VAR_GLOBAL CONSTANT   // PLC tag table "STEP7 classic symbols"
   "A" : Real := 0.5485;
   "B" : Real := 0.665E-3;
   "C" : Real := 2.805E-9;
   "A_FC343" : Real := 3.90802E-3;   // MigChange: A
   "B_FC343" : Real := -5.802000E-007;   // MigChange: B , -5.802E-7
   "C_FC343" : Real := -4.273500E-012;   // MigChange: C , -4.27350E-12
   "A_FC344" : Real := 7.64E-3;   // MigChange: A
   "B_FC344" : Real := 1.66E-5;   // MigChange: B
   "A_FC347" : Real := 3.9083E-3;   // MigChange: A
   "B_FC347" : Real := -5.775000E-007;   // MigChange: B , -5.775E-7
   "accuracy" : Real := 0.01;
END_VAR

FUNCTION "MID3" : Real   // FC96, SCL
TITLE = MID3
{ S7_Optimized_Access := 'FALSE' }
AUTHOR : hugo
FAMILY : MATH
NAME : MID3
VERSION : 1.2
// returns the mid value of 3 real inputs.
   VAR_INPUT
      in1 : Real;
      in2 : Real;
      in3 : Real;
   END_VAR
   VAR_TEMP
      tIN1 : Real;
      tIN2 : Real;
      tIN3 : Real;
   END_VAR
BEGIN


   #tIN1 := #in1;
   #tIN2 := #in2;
   #tIN3 := #in3;

   IF #tIN1 > #tIN2 THEN 
     #MID3 := #tIN1; 
     #tIN1 := #tIN2; 
     #tIN2 := #MID3; 
   END_IF;

   IF #tIN2 > #tIN3 THEN 
     #tIN2 := #tIN3; 
   END_IF;

   #MID3 := SEL(G:=#tIN1 > #tIN2, IN0:=#tIN2, IN1:=#tIN1);

   (*
   hm  1.1.2007  rev 1.1
     rewrote the function for better performance

   hm  18. mar. 2011 rev 1.2
     improve performance
   *)
END_FUNCTION

FUNCTION "MULTI_IN" : Real   // FC341, SCL
TITLE = MULTI_IN
{ S7_Optimized_Access := 'FALSE' }
AUTHOR : oscat
FAMILY : SENSOR
NAME : MULTI_IN
VERSION : 1.4
// multi_in is a signal conditioning function ehich can be configured in 8 different ways.
// it is used to read multiple sensors for the same value and protect the user from broken sensors or invalid data from sensors.
//  
// multi_in can be configured in different ways:
//     mode = 0 means the the avg of the 3 inputs is used, this mode is the default mode.
//     mode = 1 means in_1 is used.
//     mode = 2 means in_2 is used.
//     mode = 3 means in_3 is used.
//     mode = 4 means default is used.
//     mode = 5 means the lowest of the 3 external temperatures is used.
//     mode = 6 means the higest externnal temperature is used.
//     mode = 7 means the midlle input is used, if there are only two working, the lowest input is used.
//     mode > 7 ,eans output is 0 at all times.
//     in any config mode, an input higher then in_max or lower then in_min is ignored to prevent values from broken sensors or wires.
//     if all inputs are higher then in_max or lower then in_min, a default value (default) is used.
// 
// uses: MID3 [FC96]
   VAR_INPUT
      in_1 : Real;
      in_2 : Real;
      in_3 : Real;
      default : Real;
      in_min : Real;
      in_max : Real;
      mode : Int;
   END_VAR
   VAR_TEMP
      count : Int;
      F1 : Bool;
      F2 : Bool;
      F3 : Bool;
   END_VAR
BEGIN


   #F1 :=  #in_1 > #in_min AND #in_1 < #in_max;
   #F2 :=  #in_2 > #in_min AND #in_2 < #in_max;
   #F3 :=  #in_3 > #in_min AND #in_3 < #in_max;

   CASE #mode OF
   0:  #count := 0;
     IF #F1 THEN
       #count := #count + 1;
       #MULTI_IN := #in_1;
     ELSE
       #MULTI_IN := 0.0;
     END_IF;
     IF #F2 THEN
       #count := #count + 1;
       #MULTI_IN := #MULTI_IN + #in_2;
     END_IF;
     IF #F3 THEN
       #count := #count + 1;
       #MULTI_IN := #MULTI_IN + #in_3;
     END_IF;
     #MULTI_IN := SEL(G:=#count = 0, IN0:=#MULTI_IN / INT_TO_REAL(#count), IN1:=#default);

   1:  #MULTI_IN := SEL(G:=#F1, IN0:=#default, IN1:=#in_1);

   2:  #MULTI_IN := SEL(G:=#F2, IN0:=#default, IN1:=#in_2);

   3:  #MULTI_IN := SEL(G:=#F3, IN0:=#default, IN1:=#in_3);

   4:  #MULTI_IN := #default;

   5:  #MULTI_IN := SEL(G:=#F1, IN0:=#in_max, IN1:=#in_1);
     IF #F2 AND #in_2 < #MULTI_IN THEN #MULTI_IN := #in_2; END_IF;
     IF #F3 AND #in_3 < #MULTI_IN THEN #MULTI_IN := #in_3; END_IF;
     IF #MULTI_IN = #in_max THEN #MULTI_IN := #default; END_IF;

   6:  #MULTI_IN := SEL(G:=#F1, IN0:=#in_min, IN1:=#in_1);
     IF #F2 AND #in_2 > #MULTI_IN THEN #MULTI_IN := #in_2; END_IF;
     IF #F3 AND #in_3 > #MULTI_IN THEN #MULTI_IN := #in_3; END_IF;
     IF #MULTI_IN = #in_min THEN #MULTI_IN := #default; END_IF;

   7:  IF #F1 AND #F2 AND #F3 THEN #MULTI_IN := "MID3"(in1:=#in_1, in2:=#in_2, in3:=#in_3);
     ELSIF #F1 AND #F2 THEN #MULTI_IN := MIN(IN1:=#in_1, IN2:=#in_2);
     ELSIF #F1 AND #F3 THEN #MULTI_IN := MIN(IN1:=#in_1, IN2:=#in_3);
     ELSIF #F2 AND #F3 THEN #MULTI_IN := MIN(IN1:=#in_2, IN2:=#in_3);
     ELSIF #F1 THEN #MULTI_IN := #in_1;
     ELSIF #F2 THEN #MULTI_IN := #in_2;
     ELSIF #F3 THEN #MULTI_IN := #in_3;
     ELSE #MULTI_IN := #default;
     END_IF;

   END_CASE;

   (*
   hm 1.1.2007   rev 1.1
     changed midr to mid3 function

   hm  14. 10. 2008  rev 1.2
     corrected an error for in_3 overrange detection
     improved performance

   hm  11. mar. 2009 rev 1.3
     changed real constants to use dot syntax

   hm  18. jul. 2009 rev 1.4
     improved performance
   *)
END_FUNCTION

FUNCTION "RES_NI" : Real   // FC342, SCL
TITLE = RES_NI
{ S7_Optimized_Access := 'FALSE' }
AUTHOR : hugo
FAMILY : SENSOR
NAME : RES_NI
VERSION : 1.2
// this function returs the resistance for a nickel sensor for a temperature range from -60..+180 °C
   VAR_INPUT
      T : Real;
      R0 : Real;
   END_VAR
   VAR_TEMP
      T_2 : Real;
   END_VAR
BEGIN


     #T_2 := #T*#T;
     #RES_NI := #R0 + "A"*#T + "B"*#T_2 + "C"*#T_2*#T_2;


   (* revision history

   hm  4.8.2006    rev 1.0
     original version

   hm  13.9.2007    rev 1.1
     changed coding for better performance

   hm  2. dec. 2007  rev 1.2
     changed code for better performance
   *)

   (*

    Auszug aus DIN 43760 für Ni100

   °C    R    °C    R    °C  R    °C    R    °C    R

   -60   69,5   -10   94,6   40   123,0   90     154,9   140   190,9
   -55   71,9   -5     97,3   45   126,0   95     158,3   145   194,8
   -50   74,3   0     100,0   50   129,1   100   161,8   150   198,7
   -45   76,7   5     102,8   55   132,2   105   165,3   155   202,6
   -40   79,1   10     105,6   60   135,3   110   168,8   160   206,6
   -35   81,6   15     108,4   65   138,5   115   172,4   165   210,7
   -30   84,2   20     111,2   70   141,7   120   176,0   170   214,8
   -25   86,7   25     114,1   75   145,0   125   179,6   175   219,0
   -20   89,3   30     117,1   80   148,3   130   183,3   180   223,2
   -15   91,9   35     120,0   85   151,6   135   187,1        

   *)
END_FUNCTION

FUNCTION "RES_PT" : Real   // FC343, SCL
TITLE = RES_PT
{ S7_Optimized_Access := 'FALSE' }
AUTHOR : hugo
FAMILY : SENSOR
NAME : RES_PT
VERSION : 1.3
// this function returs the resistance for a platinum sensor for a temperature range from -200..+850 °C
   VAR_INPUT
      T : Real;
      R0 : Real;
   END_VAR
   VAR_TEMP
      T_2 : Real;
   END_VAR
BEGIN


   #T_2 := #T * #T;

   IF #T >= 0.0 THEN
       #RES_PT := #R0 * ( 1.0 + "A"* #T + "B_FC343" * #T_2);
   ELSE
       #RES_PT := #R0 * ( 1.0 + "A"* #T + "B_FC343" * #T_2 + "C_FC343" *(#T - 100.0) * #T_2 * #T);
   END_IF;


   (* revision history
   hm  4. aug. 2006    rev 1.1
       original version

   hm  2. dec 2007 rev 1.2
       changed code for better performance

   hm  11. mar. 2009   rev 1.3
       changed real constants to use dot syntax

   *)


   (*
    Auszug aus DIN 43760 für Pt100

   °C      R       °C      R       °C  R           °C      R           °C      R           °C      R

   -200    18,49   -100    60,25   0   100,00  100     138,50  200     175,84  300     212,02
   -195    20,65   -95     62,28   5   101,95  105     140,39  205     177,68  305     213,80
   -190    22,80   -90     64,30   10  103,90  110     142,29  210     179,51  310     215,57
   -185    24,94   -85     66,31   15  105,85  115     144,17  215     181,34  315     217,35
   -180    27,08   -80     68,33   20  107,79  120     146,06  220     183,17  320     219,12
   -175    29,20   -75     70,33   25  109,73  125     147,94  225     184,99  325     220,88
   -170    31,32   -70     72,33   30  111,67  130     149,82  230     186,82  330     222,65
   -165    33,43   -65     74,33   35  113,61   135     151,70  235     188,63  335     224,41
   -160    35,33   -60     76,33   40  115,54  140     153,58  240     190,45  340     226,17
   -155    37,63   -55     78,32   45  117,47  145     155,45  245     192,26  345     227,92
   -150    39,71   -50     80,31   50  119,40  150     157,31  250     194,07  350     229,67
   -145    41,79   -45     82,29   55  121,32  155     159,18  255     195,88  355     231,42
   -140    43,87   -40     84,27   60  123,24  160     161,04  260     197,69  360     233,17
   -135    45,94   -35     86,25   65  125,16  165     162,90  265     199,49  365     234,91
   -130    48,00  -30     88,22   70  127,07  170     164,76  270     201,29  370     236,65
   -125    50,06   -25     90,19   75  128,98  175     166,61  275     203,08  375     238,39
   -120    52,11   -20     92,16   80  130,89  180     168,46  280     204,88  380     240,13
   -115    54,15   -15     94,12   85  132,80  185     170,31  285     206,67  385     241,86
   -110    56,19   -10     96,09   90  134,70  190     172,16  290     208,45  390     243,59
   -105    58,22   -5      98,04   95  136,60  195     174,00  295     210,24  395     245,31

   *)
   (*
   revision history


   *)
END_FUNCTION

FUNCTION "RES_SI" : Real   // FC344, SCL
TITLE = RES_SI
{ S7_Optimized_Access := 'FALSE' }
AUTHOR : hugo
FAMILY : SENSOR
NAME : RES_SI
VERSION : 1.2
// this function returs the resistance for a silicon sensor for a temperature range from -50..+150 °C
// for example KTY10 normaly Rs at 25 °C
   VAR_INPUT
      T : Real;
      RS : Real;
      TS : Real;
   END_VAR
   VAR_TEMP
      TX : Real;
   END_VAR
BEGIN


   #TX := #T - #TS;
   #RES_SI := #RS * ( 1.0 + "A"* #TX + "B_FC344" * #TX * #TX);


   (* revision history
   hm  4. aug 2006 rev 1.0
       original version

   hm  2. dec 2007 rev 1.1
       changed code for better performance

   hm  11. mar. 2009   rev 1.2
       changed real constants to use dot syntax

   *)
END_FUNCTION

FUNCTION "SENSOR_INT" : Real   // FC345, SCL
TITLE = SENSOR_INT
{ S7_Optimized_Access := 'FALSE' }
AUTHOR : hugo
FAMILY : SENSOR
NAME : SENS_INT
VERSION : 1.3
// this FUNCTION calculates the REAL resistance OF a sensor RX given a parasitic resistor in parallel TO the sensor AND an additional serial resistor.
// for example a parasitic parallel resistor for a PT100 can be ignored but a series resistor is the cable to the sensor.
// for a humidity sensor, the parallel resistor is more dramatic and needs to be considered.
// the function allows to consider a parallel and serial resistor at the same time.
// with this function and known parasitic serial and parallel resistors the true resistance of the sensor can be calculated.
   VAR_INPUT
      Voltage : Real;
      Current : Real;
      RP : Real;
      RS : Real;
   END_VAR
   VAR_TEMP
      RG : Real;
   END_VAR
BEGIN


   IF #Current <> 0.0 THEN
       #RG := #Voltage / #Current;
       #SENSOR_INT := #RP * ( #RG - #RS) / ( #RP + #RS - #RG);
   END_IF;


   (* revisaion history

   hm 20.1.2007        rev 1.1
       deleted input R0 which was not needed.

   hm  2. dec 2007 rev 1.2
       corrected an error in formula and improoved speed

   hm  11. mar. 2009   rev 1.3
       changed real constants to use dot syntax

   *)
END_FUNCTION

FUNCTION "TEMP_NI" : Real   // FC346, SCL
TITLE = TEMP_NI
{ S7_Optimized_Access := 'FALSE' }
AUTHOR : hugo
FAMILY : SENSOR
NAME : TEMP_NI
VERSION : 1.5
// this function returs the temperature for a nickel sensor for a range from -60..+180 °C
   VAR_INPUT
      Res : Real;
      R0 : Real;
   END_VAR
BEGIN


   #TEMP_NI := (SQRT(0.30085225 - 2.66E-3 * (#R0 - #Res)) - 0.5485) * 751.8796992;


   (* revision history

   hm 24.1.2007        rev 1.1
       deleted unused variable A, B, C

   hm 10.9.2007        rev 1.2
       changed accuracy to 0.02 degrees to improove performace

   hm 17. 12 2007  rev 1.3
       improovements for better performance and higher accuracy

   hm  6. jan 2008 rev 1.4
       further performance improvement

   hm  10. mar. 2009   rev 1.5
       removed nested comments

   *)
END_FUNCTION

FUNCTION "TEMP_PT" : Real   // FC347, SCL
TITLE = TEMP_PT
{ S7_Optimized_Access := 'FALSE' }
AUTHOR : hugo
FAMILY : SENSOR
NAME : TEMP_PT
VERSION : 1.7
// this function returs the temperature for a platinum sensor for a range from -200..+850 °C 
// 
// uses: RES_PT [FC343]
   VAR_INPUT
      Res : Real;
      R0 : Real;
   END_VAR
   VAR_TEMP
      "step" : Real;
      X : Real;
      Y : Real;
      t1 : Real;
   END_VAR
BEGIN


   #"step" := 50.0;

   #X := "A"* #R0;
   #Y := "B_FC347" * #R0;
   IF #Res >= #R0 THEN
       #t1 := #X * #X - 4.0 * #Y * (#R0 - #Res);
       IF #t1 < 0.0 THEN
           #TEMP_PT := 10000.0;
       ELSE
           #TEMP_PT := (-#X + SQRT(#t1)) / (2.0 * #Y);
       END_IF;
   ELSE
       (* since the formula cannot be solved this is a successive approximation *)
       #TEMP_PT := -100.0;
       WHILE #"step" > "accuracy" DO
           (* test if result greater or less *)
           IF "RES_PT"(T:=#TEMP_PT,R0:=#R0) < #Res THEN #TEMP_PT := #TEMP_PT + #"step"; ELSE #TEMP_PT := #TEMP_PT - #"step"; END_IF;
           (* pt^ := pt^ - 8388608; *)  (* this is a super fast divide by 2 method for non floating point CPUs *)
           (* the alternative code: step := step * 0.5; *)
           #"step" := #"step" * 0.5;
       END_WHILE;
   END_IF;

   (* revision history

   rev 1.1 hm 24.1.2007    
       deleted unused variable C

   rev 1.2 hm 10.9.2007
       reduced accuracy to 0.02 to shorten execution time

   rev 1.3 hm  2. dec 2007
       changed code for better performance

   rev 1.4 hm  23. dec 2007
       avoid a negative square root if input values are wrong

   rev 1.5 hm 5. jan 2008
       replaced / 2 with * 0.5 for better performance

   hm  31. oct. 2008   rev 1.6
       improved performance

   hm  11. mar. 2009   rev 1.7
       changed real constants to use dot syntax

   *)
END_FUNCTION

FUNCTION "TEMP_SI" : Real   // FC348, SCL
TITLE = TEMP_SI
{ S7_Optimized_Access := 'FALSE' }
AUTHOR : hugo
FAMILY : SENSOR
NAME : TEMP_SI
VERSION : 1.5
// this function returs the temperature for a silicon sensor for a range from -50..+150 °C
// for example KTY10 RS at TS normally 25 °C
   VAR_INPUT
      Res : Real;
      RS : Real;
      TS : Real;
   END_VAR
BEGIN


   #TEMP_SI := (-7.64E-3 + SQRT(#Res/#RS* 6.64E-5 - 0.803E-5)) * 30120.48193 + #TS;


   (* revision history

   hm 24.1.2007        rev 1.1
       the function would only work for TS = 25, now it works for other values of ts.

   hm 10.9.2007        rev 1.2
       changed the function to use successive approcimation to avoid an error generated by a sqrt from a negative result.
       changed accuracy to 0.02 degrees to shorten execution time

   hm 17. 12 2007  rev 1.3
       improovements for better performance

   hm  6. jan 2008 rev 1.4
       further performance improvement

   hm  10. mar. 2009   rev 1.5
       removed nested comments

   *)
END_FUNCTION

FUNCTION "TEMP_NTC" : Real   // FC411, SCL
TITLE = TEMP_NTC
{ S7_Optimized_Access := 'FALSE' }
AUTHOR : hugo
FAMILY : SENSOR
NAME : TEMP_NTC
VERSION : 1.1
// this function returs the temperature for a NTC sensor for a range from 0..85 °C.
// RN is the resistance at 25 °C and B is a constant for the given sensor.
   VAR_INPUT
      RES : Real;
      RN : Real;
      "B" : Real;
   END_VAR
BEGIN


   IF #RES > 0.0 THEN
       #TEMP_NTC := #"B" * 298.15 / (#"B" + LN(#RES / #RN) * 298.15) -273.15;
   END_IF;


   (* revision history

   hm 30. dec. 2008    rev 1.0
       original version

   hm  11. mar. 2009   rev 1.1
       changed real constants to use dot syntax

   *)
END_FUNCTION

FUNCTION "RES_NTC" : Real   // FC412, SCL
TITLE = RES_NTC
{ S7_Optimized_Access := 'FALSE' }
AUTHOR : hugo
FAMILY : SENSOR
NAME : RES_NTC
VERSION : 1.1
// this function returs the resistance for a NTC sensor for a given temperature in °C.
// RN is the resistance at 25 °C and B is a constant for the given sensor.
   VAR_INPUT
      T : Real;
      RN : Real;
      "B" : Real;
   END_VAR
BEGIN


   #RES_NTC := #RN * EXP(#"B" * (1.0 / (#T+273.15) - 0.00335401643468053));


   (* revision history

   hm 30. dec. 2008    rev 1.0
       original version

   hm  11. mar. 2009   rev 1.1
       changed real constants to use dot syntax

   *)
END_FUNCTION

// ===== PLC "List Processing"  Unspecific CPU S7 300 =====

DATA_BLOCK "TEMP"   // DB7
TITLE = temporary Strings
{ S7_Optimized_Access := 'FALSE' }
AUTHOR : dalbi
FAMILY : xS7
NAME : DBTEMP
VERSION : 1.1
   VAR
      STR1 : String[254];
      STR2 : String[254];
      STR3 : String[254];
      TEMP : String[254];
   END_VAR
BEGIN
END_DATA_BLOCK

FUNCTION_BLOCK "LIST_NEXT"   // FB231, SCL
TITLE = LIST_NEXT
{ S7_Optimized_Access := 'FALSE' }
AUTHOR : hugo
FAMILY : LISTPRO
NAME : LNEXT
VERSION : 2.0
// LIST_NEXT retrieves the next element of a list, starting from element 1 after reset or first init.
// when the end of the lisat is reached a '' empty string is returned and NUL is set to true.
// die liste liegt als string von elementen vor die mit den zeichen SEP am anfang markiert sind.
   VAR_INPUT
      SEP : Byte;
      RST : Bool;
   END_VAR
   VAR_OUTPUT
      LEL : String[254];
      po AT LEL : Struct
         length : Byte;
         act_length : Byte;
         str : Array[1..254] of Byte;
      END_STRUCT;
      NUL : Bool;
   END_VAR
   VAR_IN_OUT
      LIST : String[254];
      pt AT LIST : Struct
         length : Byte;
         act_length : Byte;
         str : Array[1..254] of Byte;
      END_STRUCT;
   END_VAR
   VAR
      pos : Int := 1;
      c : Byte;
      write : Int;
   END_VAR
BEGIN


   //pt := ADR(LIST);
   //po := ADR(LEL);

   IF #RST THEN
     #pos := 1;
   END_IF;

   IF #pt.str[#pos] = 0 OR #pos = BYTE_TO_INT(#pt.act_length) THEN
     #LEL := '';
     #NUL := TRUE;
   ELSE
     #NUL := FALSE;
     #write := 1;
     FOR #pos := #pos + 1 TO BYTE_TO_INT(#pt.act_length) DO
       #c := #pt.str[#pos];
       IF #c = 0 OR #c = #SEP THEN
         #po.str[#write] := 0;
         RETURN;
       ELSE
         #po.str[#write] := #pt.str[#pos];
         #write := #write + 1;
       END_IF;
     END_FOR;
   END_IF;

   #po.length := #pt.length;
   #po.act_length := INT_TO_BYTE(#write);


   (* revision histroy
   hm  25. jun. 2008 rev 1.0
     original release

   hm  19. jan. 2011 rev 1.1
     changed string(255) to string(LIST_LENGTH)  

   hm  21. mar. 2011 rev 2.0
     all elements start with SEP

   *)
END_FUNCTION_BLOCK

FUNCTION "CHR_TO_STRING" : String[254]   // FC227, SCL
TITLE = CHR_TO_STRING
{ S7_Optimized_Access := 'FALSE' }
AUTHOR : hugo
FAMILY : STRINGS
NAME : CHRSTR
VERSION : 1.3
// CHR creates a character from a byte input and stuffs it in a one character length string.
   VAR_INPUT
      C : Byte;
   END_VAR
   VAR_TEMP
      tCHR : String[1];
      _CHR AT tCHR : Array[0..2] of Byte;
   END_VAR
BEGIN


   #_CHR[0] := 1;   (* length *)
   #_CHR[1] := 1;   (* actual length *)
   #_CHR[2] := #C; 
   #CHR_TO_STRING := #tCHR;

   (* revision history
   hm  16 jan 2007     rev 1.0
       original version

   hm  4. feb. 2008    rev 1.1
       return string would not be terminated properly

   hm  29. mar. 2008   rev 1.2
       changed STRING to STRING(1)

   hm  17. dec. 2008   rev 1.3
       changed name of function from chr to chr_to_string
   *)
END_FUNCTION

FUNCTION "LIST_CLEAN" : Bool   // FC389, SCL
TITLE = LIST_CLEAN
{ S7_Optimized_Access := 'FALSE' }
AUTHOR : hugo
FAMILY : LISTPRO
NAME : LCLEAN
VERSION : 2.0
// LIST_CLEAN bereinigt eine liste von leeren Elementen.
// die liste liegt als string von elementen vor die mit den zeichen SEP am anfang markiert sind.
   VAR_INPUT
      SEP : Byte;
   END_VAR
   VAR_IN_OUT
      LIST : String[254];
      pt AT LIST : Struct
         length : Byte;
         act_length : Byte;
         str : Array[1..254] of Byte;
      END_STRUCT;
   END_VAR
   VAR_TEMP
      read : Int;
      write : Int;
      last : Byte;
      c : Byte;
   END_VAR
BEGIN


   #read := 1;
   #write := 1;

   FOR #read := 1 TO BYTE_TO_INT(#pt.act_length) DO //LIST_LENGTH = 254
     #c := #pt.str[#read];               (* read character from list *)
     IF #c = 0 THEN EXIT;           (* exit the loop if character definbes end of string *)
     ELSIF #c <> #SEP OR #SEP <> #last THEN  (* copy element from read to write position unless a double sep character is present *)
       #pt.str[#write] := #c;
       #write := #write + 1;
     END_IF;
     #last := #c;                  (* remember last character *)
   END_FOR;

   IF #last = #SEP THEN #write := #write - 1; END_IF;    (* if last character is sep then delete empty element at end *)
   IF #write <= BYTE_TO_INT(#pt.act_length) THEN #pt.str[#write] := 0;  END_IF;    (* terminate string with 0 *)

   #LIST_CLEAN := TRUE;           (* retrun TRUE *)


   (* revision histroy
   hm  28. jun. 2008 rev 1.0
     original release

   hm  19. jan. 2011 rev 1.1
     changed string(255) to string(LIST_LENGTH)

   hm  21. mar. 2011 rev 2.0
     all elements start with SEP

   *)
END_FUNCTION

FUNCTION "LIST_GET" : String[254]   // FC390, SCL
TITLE = LIST_GET
{ S7_Optimized_Access := 'FALSE' }
AUTHOR : hugo
FAMILY : LISTPRO
NAME : LGET
VERSION : 2.0
// LIST_GET liefert das element an der stelle pos einer liste.
// die liste liegt als string von elementen vor die mit den zeichen SEP am anfang makiert sind.
   VAR_INPUT
      SEP : Byte;
      POS : Int;
   END_VAR
   VAR_IN_OUT
      LIST : String[254];
      pt AT LIST : Struct
         length : Byte;
         act_length : Byte;
         str : Array[1..254] of Byte;
      END_STRUCT;
   END_VAR
   VAR_TEMP
      tLIST_GET : String[254];
      po AT tLIST_GET : Struct
         length : Byte;
         act_length : Byte;
         str : Array[1..254] of Byte;
      END_STRUCT;
      i : Int;
      o : Int;
      cnt : Int;
      c : Byte;
   END_VAR
BEGIN


   #i := 1;
   #o := 1;
   #cnt := 0;

   REPEAT
     #c := #pt.str[#i];
     IF #cnt = #POS THEN           (* copy element to output string *)
       IF #c = #SEP  THEN EXIT; END_IF;    (* next element stop copy and finish *)
       #po.str[#o] := #c;
       #o := #o + 1;
     ELSIF #c = #SEP THEN
       #cnt := #cnt + 1;
     END_IF;
     #i := #i + 1;
   UNTIL
     (#i = BYTE_TO_INT(#pt.act_length)) OR (#c = 0)
   END_REPEAT;
   #po.act_length := INT_TO_BYTE(#o);            (* close the output string *)
   #po.length := #pt.length;

   #LIST_GET := #tLIST_GET;


   (* revision histroy
   hm  20. jun. 2008 rev 1.0
     original release

   hm  19. jan. 2011 rev 1.1
     changed string(255) to strring(LIST_LENGTH)

   hm  21. mar. 2011 rev 2.0
     all list elements start with SEP
   *)
END_FUNCTION

FUNCTION "LIST_INSERT" : Bool   // FC391, SCL
TITLE = LIST_INSERT
{ S7_Optimized_Access := 'FALSE' }
AUTHOR : hugo
FAMILY : LISTPRO
NAME : LINS
VERSION : 2.0
// LIST_INSERT setzt ein element an der stelle pos in eine liste ein.
// die liste liegt als string von elementen vor die mit den zeichen SEP am anfang markiert sind.
// 
// uses: CONCAT [FC2]
//       CHR_TO_STRING [FC227]
//       INSERT [FC17]
//       LEN [FC21]
//       TEMP [DB7]
   VAR_INPUT
      SEP : Byte;
      POS : Int;
      INS : String[254];
      _INS AT INS : Struct
         length : Byte;
         act_length : Byte;
         str : Array[1..254] of Byte;
      END_STRUCT;
   END_VAR
   VAR_IN_OUT
      LIST : String[254];
      pt AT LIST : Struct
         length : Byte;
         act_length : Byte;
         str : Array[1..254] of Byte;
      END_STRUCT;
   END_VAR
   VAR_TEMP
      read : Int;
      cnt : Int;
      sx : String[1];
   END_VAR
BEGIN


   #read := 1;
   #cnt := 1;

   "TEMP".STR1 := #LIST;
   "TEMP".STR2 := #INS;

   IF LEN("TEMP".STR2) + 1 + LEN("TEMP".STR1) > BYTE_TO_INT(#pt.length) THEN
     #LIST_INSERT := FALSE;
   ELSE
     #LIST_INSERT := TRUE;
     (* search for position *)
     WHILE #read < BYTE_TO_INT(#pt.length) DO
       IF #cnt >= #POS THEN
         #sx := "CHR_TO_STRING"(#SEP);
         "TEMP".STR2 := CONCAT(IN1:=#sx,IN2:="TEMP".STR2);
         "TEMP".STR1 := INSERT(IN1:="TEMP".STR1,IN2:="TEMP".STR2,P:=#read - 1);
         #LIST_INSERT := TRUE;
         RETURN;
       END_IF;
       #LIST := "TEMP".STR1;
       IF #pt.str[#read]  = 0 THEN        (* list is too short add empty element *)
         #pt.str[#read] := #SEP;
         #pt.str[#read + 1] := 0;
       END_IF;
       #read := #read + 1;
       IF #pt.str[#read] = #SEP OR #pt.str[#read] = 0 THEN #cnt := #cnt + 1; END_IF;
     END_WHILE;
   END_IF;



   (* revision histroy
   hm  28. jun. 2008 rev 1.0
     original release

   hm  17. dec. 2008 rev 1.1
     changes name of function chr to chr_to_string

   hm  19. jan. 2011 rev 1.2
     changed string(255) to string(LIST_LENGTH)

   hm  21. mar. 2011 rev 2.0
     all list elements start with SEP

   *)
END_FUNCTION

FUNCTION "LIST_LEN" : Int   // FC392, SCL
TITLE = LIST_LEN
{ S7_Optimized_Access := 'FALSE' }
AUTHOR : hugo
FAMILY : LISTPRO
NAME : LLEN
VERSION : 2.0
// LIST_LEN liefert die anzahl der elemente einer liste.
// die liste liegt als string von elementen vor die mit den zeichen SEP am anfang markiert sind.
   VAR_INPUT
      SEP : Byte;
   END_VAR
   VAR_IN_OUT
      LIST : String[254];
      pt AT LIST : Struct
         length : Byte;
         act_length : Byte;
         str : Array[1..254] of Byte;
      END_STRUCT;
   END_VAR
   VAR_TEMP
      l : Int;
      pos : Int;
      c : Byte;
   END_VAR
BEGIN


   //pt := ADR(LIST);
   #pos := 1;
   #LIST_LEN := 0;
   REPEAT
     #c := #pt.str[#pos];
     IF #c = #SEP THEN #LIST_LEN := #LIST_LEN + 1; END_IF;
     #pos := #pos + 1;
   UNTIL
     #c = 0 OR #pos > BYTE_TO_INT(#pt.act_length)  //LIST_LENGTH
   END_REPEAT;


   (* revision histroy
   hm  25. jun. 2008 rev 1.0
     original release

   hm  16. oct. 2008 rev 1.1
     fixed a problem where list_len would only work up to LIST_LENGTH

   hm  19. jan. 2001 rev 1.2
     changed string(255) to string(LIST_LENGTH)

   hm  21. mar. 2011 rev 2.0
     all list elements start with SEP

   *)
END_FUNCTION

FUNCTION "LIST_ADD" : Bool   // FC393, SCL
TITLE = LIST_ADD
{ S7_Optimized_Access := 'FALSE' }
AUTHOR : hugo
FAMILY : LISTPRO
NAME : LISTADD
VERSION : 2.0
// LIST_ADD hängt ein weiteres element ans ende einer liste.
// die liste liegt als string von elementen vor die mit den zeichen SEP am anfang makiert sind.
// 
// uses: CONCAT [FC2]
//       CHR_TO_STRING [FC227]
//       LEN [FC21]
//       TEMP [DB7]
   VAR_INPUT
      SEP : Byte;
   END_VAR
   VAR_IN_OUT
      INS : String[254];
      LIST : String[254];
      tLIST AT LIST : Struct
         length : Byte;
         act_length : Byte;
         str : Array[1..254] of Byte;
      END_STRUCT;
   END_VAR
   VAR_TEMP
      sx : String[1];
   END_VAR
BEGIN


   "TEMP".STR1 := #INS;
   "TEMP".STR2 := #LIST;

   #sx := "CHR_TO_STRING"(#SEP);     (* convert separation character to string *)
   "TEMP".STR1 := CONCAT(IN1:=#sx,IN2:="TEMP".STR1);         (* start element with separation character *)

   IF LEN("TEMP".STR2) + LEN("TEMP".STR1) > BYTE_TO_INT(#tLIST.length) THEN
     #LIST_ADD := FALSE;          (* return false if element does not fit *)
   ELSE
     "TEMP".STR2 := CONCAT(IN1:="TEMP".STR2,IN2:="TEMP".STR1);
     #LIST_ADD := TRUE;
   END_IF;

   #LIST := "TEMP".STR2;

   (* revision histroy

   hm  21. mar. 2011 rev 2.0
     original release
   *)
END_FUNCTION

FUNCTION "LIST_RETRIEVE_LAST" : String[254]   // FC395, SCL
TITLE = LIST_RETRIEVE_LAST
{ S7_Optimized_Access := 'FALSE' }
AUTHOR : hugo
FAMILY : LISTPRO
NAME : LRETLA
VERSION : 2.0
// LIST_RETRIEVE_LAST liefert das letzte element einer liste und löscht das element aus der liste.
// die liste liegt als string von elementen vor die mit den zeichen SEP beginnen.
// 
// uses: MID [FC26]
//       TEMP [DB7]
   VAR_INPUT
      SEP : Byte;
   END_VAR
   VAR_IN_OUT
      LIST : String[254];
      pt AT LIST : Struct
         length : Byte;
         act_length : Byte;
         str : Array[1..254] of Byte;
      END_STRUCT;
   END_VAR
   VAR_TEMP
      i : Int;
      last : Int;
      c : Byte;
   END_VAR
BEGIN


   "TEMP".STR1 := #LIST;
   #LIST_RETRIEVE_LAST := '';
   #last := 1;

   (* search position of last element *)
   FOR #i := 1 TO BYTE_TO_INT(#pt.act_length) DO
     #c := #pt.str[#i];
     IF #c = 0 THEN
       EXIT;
     ELSIF #c = #SEP THEN
       #last := #i;
     END_IF;
   END_FOR;
   (* return last element of list *)
   "TEMP".STR2 := MID(IN:="TEMP".STR1,L:=BYTE_TO_INT(#pt.act_length),P:=#last + 1);

   #LIST_RETRIEVE_LAST := "TEMP".STR2;


   (* revision histroy
   hm  21. mar. 2011 rev 2.0
     new module
   *)
END_FUNCTION

FUNCTION "LIST_RETRIEVE" : String[254]   // FC406, SCL
TITLE = LIST_RETRIEVE
{ S7_Optimized_Access := 'FALSE' }
AUTHOR : hugo
FAMILY : LISTPRO
NAME : LRETR
VERSION : 2.0
// LIST_RETRIEVE liefert das element an der stelle pos einer liste und löscht das element aus der liste.
// die liste liegt als string von elementen vor die mit den zeichen SEP separiert sind.
   VAR_INPUT
      SEP : Byte;
      POS : Int;
   END_VAR
   VAR_IN_OUT
      LIST : String[254];
      pt AT LIST : Struct
         length : Byte;
         act_length : Byte;
         str : Array[1..254] of Byte;
      END_STRUCT;
   END_VAR
   VAR_TEMP
      i : Int;
      o : Int;
      w : Int;
      cnt : Int;
      c : Byte;
      tLIST_RETRIEVE : String[254];
      po AT tLIST_RETRIEVE : Struct
         length : Byte;
         act_length : Byte;
         str : Array[1..254] of Byte;
      END_STRUCT;
   END_VAR
BEGIN


   #po.act_length := #pt.act_length;
   #po.length := #pt.length;

   #o := 1;
   #w := 1;
   #cnt := 0;

   IF #POS > 0 THEN
     FOR #i := 1 TO BYTE_TO_INT(#pt.act_length) DO
       #c := #pt.str[#i];
       IF #c = 0 THEN
         #po.str[#o] := 0;
         IF #cnt < #POS THEN #pt.str[#w + 1] := 0; ELSE #pt.str[#w] := 0; END_IF;
         RETURN;
       ELSIF #cnt = #POS AND #c <> #SEP THEN       (* we have found the element *)
         #po.str[#o] := #pt.str[#i];
         #o := #o + 1;
       ELSIF #cnt >= #POS THEN
         #pt.str[#w] := #c;
         #w := #w + 1;
       ELSE
         #w := #i;
       END_IF;
       IF #c = #SEP THEN #cnt := #cnt + 1; END_IF;
     END_FOR;
   ELSE
     #LIST_RETRIEVE := '';
   END_IF;


   (* revision histroy
   hm  28. jun. 2008 rev 1.0
     original release

   hm  19. jan. 2011 rev 1.1
     changed string(255) to string(LIST_LENGTH)

   hm  21. mar. 2011 rev 2.0
     all elements start with SEP
   *)
END_FUNCTION

// ===== PLC "Logic FF edge triggered"  Unspecific CPU S7 300 =====

FUNCTION_BLOCK "COUNT_BR"   // FB77, SCL
TITLE = COUNT_BR
{ S7_Optimized_Access := 'FALSE' }
AUTHOR : hugo
FAMILY : FFETRIG
NAME : COUNT_BR
VERSION : 1.0
// Count_R is a byte counter with independen up and dn inputs. the counter counts from 0 to mx and continues at 0 after is has reached mx
// a step input sets the counters stepping width.
// 
// uses: INC [FC90]
   VAR_INPUT
      SET : Bool;
      IN : Byte;
      UP : Bool;
      DN : Bool;
      "STEP" : Byte := B#16#1;
      MX : Byte := B#16#FF;
      RST : Bool;
   END_VAR
   VAR_OUTPUT
      CNT : Byte;
   END_VAR
   VAR
      last_up : Bool;
      last_dn : Bool;
   END_VAR
BEGIN


     IF #RST THEN
       #CNT := 0;
     ELSIF #SET THEN
       #CNT := INT_TO_BYTE(LIMIT(MN:=0,IN:=BYTE_TO_INT(#IN),MX:=BYTE_TO_INT(#MX)));
     ELSIF #UP AND NOT #last_up THEN
       #CNT := INT_TO_BYTE("INC"(X:=BYTE_TO_INT(#CNT),D:=BYTE_TO_INT(#"STEP"),M:=BYTE_TO_INT(#MX)));
     ELSIF #DN AND NOT #last_dn THEN
       #CNT := INT_TO_BYTE("INC"(X:=BYTE_TO_INT(#CNT),D:=-BYTE_TO_INT(#"STEP"),M:=BYTE_TO_INT(#MX)));
     END_IF;
     #last_up := #UP;
     #last_dn := #DN;

   (* revision history
   hm  16. jan 2008  rev 1.0
     original version

   *)
END_FUNCTION_BLOCK

FUNCTION_BLOCK "COUNT_DR"   // FB78, SCL
TITLE = COUNT_DR
{ S7_Optimized_Access := 'FALSE' }
AUTHOR : hugo
FAMILY : FFETRIG
NAME : COUNT_DR
VERSION : 1.1
// Count_DR is a DWORD counter with independen up and dn inputs. the counter counts from 0 to mx and continues at 0 after is has reached mx
// a step input sets the counters stepping width.
   VAR_INPUT
      SET : Bool;
      IN : DWord;
      UP : Bool;
      DN : Bool;
      "STEP" : DWord := DW#16#1;
      MX : DWord := DW#16#FFFFFFFF;
      RST : Bool;
   END_VAR
   VAR_OUTPUT
      CNT : DWord;
   END_VAR
   VAR
      last_up : Bool;
      last_dn : Bool;
   END_VAR
BEGIN


   IF #RST THEN
     #CNT := 0;
   ELSIF #SET THEN
     #CNT := DINT_TO_DWORD(LIMIT(MN:=0,IN:=DWORD_TO_DINT(#IN),MX:=DWORD_TO_DINT(#MX)));
   ELSIF #UP AND NOT #last_up THEN
     IF DWORD_TO_DINT(#"STEP") > DWORD_TO_DINT(#MX) - DWORD_TO_DINT(#CNT) THEN
         #CNT := DINT_TO_DWORD(DWORD_TO_DINT(#CNT) - DWORD_TO_DINT(#MX) + DWORD_TO_DINT(#"STEP") - 1);
     ELSE
         #CNT := DINT_TO_DWORD(DWORD_TO_DINT(#CNT) + DWORD_TO_DINT(#"STEP"));
     END_IF;
   ELSIF #DN AND NOT #last_dn THEN
     IF DWORD_TO_DINT(#"STEP") > DWORD_TO_DINT(#CNT) THEN
         #CNT := DINT_TO_DWORD(DWORD_TO_DINT(#CNT) - DWORD_TO_DINT(#"STEP") + DWORD_TO_DINT(#MX) + 1);
     ELSE
         #CNT := DINT_TO_DWORD(DWORD_TO_DINT(#CNT) - DWORD_TO_DINT(#"STEP"));
     END_IF;
   END_IF;
   #last_up := #UP;
   #last_dn := #DN;


   (* revision history
   hm  12. jun 2008  rev 1.0
     original version

   hm  20. jan. 2011 rev 1.1
     corrected init value of MX to 16#FFFFFFFF

   *)
END_FUNCTION_BLOCK

FUNCTION_BLOCK "FF_D2E"   // FB79, SCL
TITLE = FF_D2E
{ S7_Optimized_Access := 'FALSE' }
AUTHOR : hugo
FAMILY : FFETRIG
NAME : FF_D2E
VERSION : 1.3
// dual D-type flip flop with reset and rising clock trigger
   VAR_INPUT
      D0 : Bool;
      D1 : Bool;
      CLK : Bool;
      RST : Bool;
   END_VAR
   VAR_OUTPUT
      Q0 : Bool;
      Q1 : Bool;
   END_VAR
   VAR
      edge : Bool;
   END_VAR
BEGIN


   IF #RST THEN
       #Q0 := FALSE;
       #Q1 := FALSE;
   ELSIF #CLK AND NOT #edge THEN
       #Q0 := #D0;
       #Q1 := #D1;
   END_IF;
   #edge := #CLK;


   (* revision history
   hm  25. dec 2007    rev 1.0
       original version

   hm  27. dec 2007    rev 1.1
       changed code for better performance

   hm  30. oct. 200    rev 1.2
       deleted unnecessary init with 0

   hm  14. mar. 2009   rev 1.3
       removed double assignments

   *)
END_FUNCTION_BLOCK

FUNCTION_BLOCK "FF_D4E"   // FB80, SCL
TITLE = FF_D4E
{ S7_Optimized_Access := 'FALSE' }
AUTHOR : hugo
FAMILY : FFETRIG
NAME : FF_D4E
VERSION : 1.3
// quad D-type flip flop with reset and rising clock trigger
   VAR_INPUT
      D0 : Bool;
      D1 : Bool;
      D2 : Bool;
      D3 : Bool;
      CLK : Bool;
      RST : Bool;
   END_VAR
   VAR_OUTPUT
      Q0 : Bool;
      Q1 : Bool;
      Q2 : Bool;
      Q3 : Bool;
   END_VAR
   VAR
      edge : Bool;
   END_VAR
BEGIN


   IF #RST THEN
       #Q0 := FALSE;
       #Q1 := FALSE;
       #Q2 := FALSE;
       #Q3 := FALSE;
   ELSIF #CLK AND NOT #edge THEN
       #Q0 := #D0;
       #Q1 := #D1;
       #Q2 := #D2;
       #Q3 := #D3;
   END_IF;
   #edge := #CLK;


   (* revision history
   hm  4. aug 2006 rev 1.0
       original version

   hm  27. dec 2007    rev 1.1
       changed code for better performance

   hm  30. oct. 200    rev 1.2
       deleted unnecessary init with 0

   hm  14. mar. 2009   rev 1.3
       removed double assignments

   *)
END_FUNCTION_BLOCK

FUNCTION_BLOCK "FF_DRE"   // FB81, SCL
TITLE = FF_DRE
{ S7_Optimized_Access := 'FALSE' }
AUTHOR : hugo
FAMILY : FFETRIG
NAME : FF_DRE
VERSION : 1.2
// D-type flip flop with set, reset and rising clock trigger
   VAR_INPUT
      SET : Bool;
      D : Bool;
      CLK : Bool;
      RST : Bool;
   END_VAR
   VAR_OUTPUT
      Q : Bool;
   END_VAR
   VAR
      edge : Bool;
   END_VAR
BEGIN


   IF #RST OR #SET THEN
       #Q := NOT #RST;
   ELSIF #CLK AND NOT #edge THEN
       #Q := #D;
   END_IF;
   #edge := #CLK;

   (* revision history
   hm  4. aug 2006     rev 1.0
       original version

   hm  27. dec 2007    rev 1.1
       changed code for better performance

   hm  30. oct. 2008   rev 1.2
       optimized performance
   *)
END_FUNCTION_BLOCK

FUNCTION_BLOCK "FF_JKE"   // FB82, SCL
TITLE = FF_JKE
{ S7_Optimized_Access := 'FALSE' }
AUTHOR : hugo
FAMILY : FFETRIG
NAME : FF_JKE
VERSION : 1.2
// JK-type flip flop with set, reset and rising clock trigger
// set and reset are asynchron while the FF is rising edge triggered
// J=0 and K=0 and CLK >>> no action
// J=1 and K=0 and CLK >>> output = 1
// J=0 and K=1 and CLK >>> output = 0
// J=1 and K=1 and CLK >>> toggle output
   VAR_INPUT
      SET : Bool;
      J : Bool;
      CLK : Bool;
      K : Bool;
      RST : Bool;
   END_VAR
   VAR_OUTPUT
      Q : Bool;
   END_VAR
   VAR
      edge : Bool;
   END_VAR
BEGIN


   IF #RST OR #SET THEN
       #Q := NOT #RST;
   ELSIF #CLK AND NOT #edge THEN
       IF #J XOR #K THEN #Q := #J;
       ELSE #Q := #K XOR #Q;
       END_IF;
   END_IF;
   #edge := #CLK;

   (* revision history
   hm  4. aug 2006     rev 1.0
       original version

   hm  27. dec 2007    rev 1.1
       changed code for better performance

   hm  30. oct. 2008   rev 1.2
       optimized performance
   *)
END_FUNCTION_BLOCK

FUNCTION_BLOCK "FF_RSE"   // FB83, SCL
TITLE = FF_RSE
{ S7_Optimized_Access := 'FALSE' }
AUTHOR : hugo
FAMILY : FFETRIG
NAME : FF_RSE
VERSION : 1.0
// this is a rising edge triggered rs flip flop
// a rising edge on CS sets Q = TRUE and a rising edge on CR sets Q = FALSE.
// CR has priority over CS.
   VAR_INPUT
      CS : Bool;
      CR : Bool;
      RST : Bool;
   END_VAR
   VAR_OUTPUT
      Q : Bool;
   END_VAR
   VAR
      es : Bool;
      er : Bool;
   END_VAR
BEGIN


   IF #RST THEN
       (* asynchronous reset *)
       #Q := FALSE;
   ELSIF #CR AND NOT #er THEN
       (* rising edge on CR *)
       #Q := FALSE;
   ELSIF #CS AND NOT #es THEN
       (* rising edge on CS *)
       #Q := TRUE;
   END_IF;

   #es := #CS;
   #er := #CR;

   (* revision history

   hm  16. jul. 2008   rev 1.0
       original version

   *)
END_FUNCTION_BLOCK

FUNCTION_BLOCK "SELECT_8"   // FB84, SCL
TITLE = SELECT_8
{ S7_Optimized_Access := 'FALSE' }
AUTHOR : hugo
FAMILY : FFETRIG
NAME : SELECT8
VERSION : 1.1
// select_8 selects one of 8 outputs at any time. the outputscan be selected by up or down keys and an independent anable switches all outouts off if set false
// 
// uses: INC [FC90]
   VAR_INPUT
      "E" : Bool;
      SET : Bool;
      IN : Byte;
      UP : Bool;
      DN : Bool;
      RST : Bool;
   END_VAR
   VAR_OUTPUT
      Q0 : Bool;
      Q1 : Bool;
      Q2 : Bool;
      Q3 : Bool;
      Q4 : Bool;
      Q5 : Bool;
      Q6 : Bool;
      Q7 : Bool;
      STATE : Int;
   END_VAR
   VAR
      last_up : Bool;
      last_dn : Bool;
   END_VAR
BEGIN


   IF #RST THEN
       #STATE := 0;
   ELSIF #SET THEN
       #STATE := BYTE_TO_INT(#IN);
   ELSIF #UP AND NOT #last_up THEN
       #STATE := "INC"(X:=#STATE,D:=1,M:=7);
   ELSIF #DN AND NOT #last_dn THEN
       #STATE := "INC"(X:=#STATE,D:=-1,M:=7);
   END_IF;
   #last_up := #UP;
   #last_dn := #DN;

   #Q0 := FALSE;
   #Q1 := FALSE;
   #Q2 := FALSE;
   #Q3 := FALSE;
   #Q4 := FALSE;
   #Q5 := FALSE;
   #Q6 := FALSE;
   #Q7 := FALSE;

   IF #"E" THEN
       CASE #STATE OF
         0: #Q0 := TRUE;
         1: #Q1 := TRUE;
         2: #Q2 := TRUE;
         3: #Q3 := TRUE;
         4: #Q4 := TRUE;
         5: #Q5 := TRUE;
         6: #Q6 := TRUE;
         7: #Q7 := TRUE;
       END_CASE;
   END_IF;


   (* revision history
   hm  16. jan 2008    rev 1.0
       original version

   hm  27. feb. 2009   rev 1.1
       renamed input en to e
   *)
END_FUNCTION_BLOCK

FUNCTION_BLOCK "SHR_4E"   // FB87, SCL
TITLE = SHR_4E
{ S7_Optimized_Access := 'FALSE' }
AUTHOR : hugo
FAMILY : FFETRIG
NAME : SHR_4E
VERSION : 1.1
// 4 bit shift register with reset
   VAR_INPUT
      SET : Bool;
      D0 : Bool;
      CLK : Bool;
      RST : Bool;
   END_VAR
   VAR_OUTPUT
      Q0 : Bool;
      Q1 : Bool;
      Q2 : Bool;
      Q3 : Bool;
   END_VAR
   VAR
      "m" : Bool;
   END_VAR
BEGIN


   (* trig.Q signals a rising edge on clk *)
   (* trig(clk := clk); *)

   IF #SET OR #RST THEN
       #Q0 := NOT #RST;
       #Q1 := NOT #RST;
       #Q2 := NOT #RST;
       #Q3 := NOT #RST;
   ELSIF #CLK AND NOT #"m" THEN    //ELSIF trig.Q THEN
       #Q3 := #Q2;
       #Q2 := #Q1;
       #Q1 := #Q0;
       #Q0 := #D0;
   END_IF;

   #"m" := #CLK;


   (* revision history
   hm  4. aug. 2006    rev 1.0
       original version

   hm  25. oct. 2008   rev 1.1
       optimized code

   *)
END_FUNCTION_BLOCK

FUNCTION_BLOCK "SHR_4UDE"   // FB88, SCL
TITLE = SHR_4UDE
{ S7_Optimized_Access := 'FALSE' }
AUTHOR : hugo
FAMILY : FFETRIG
NAME : SHR4UDE
VERSION : 1.2
// 4 bit shift register with reset up / down direction input
   VAR_INPUT
      SET : Bool;
      D0 : Bool;
      D3 : Bool;
      CLK : Bool;
      DN : Bool;
      RST : Bool;
   END_VAR
   VAR_OUTPUT
      Q0 : Bool;
      Q1 : Bool;
      Q2 : Bool;
      Q3 : Bool;
   END_VAR
   VAR
      "m" : Bool;
   END_VAR
BEGIN


   (* trig.Q signals a rising edge on clk *)
   (* trig(clk := clk); *)

   IF #SET OR #RST THEN
       #Q0 := NOT #RST;
       #Q1 := #Q0;
       #Q2 := #Q0;
       #Q3 := #Q0;
   ELSIF #CLK AND NOT #"m" THEN
       IF #DN THEN
           #Q0 := #Q1;
           #Q1 := #Q2;
           #Q2 := #Q3;
           #Q3 := #D3;
       ELSE
           #Q3 := #Q2;
           #Q2 := #Q1;
           #Q1 := #Q0;
           #Q0 := #D0;
       END_IF;
   END_IF;

   #"m" := #CLK;


   (* revision history
   hm  4. aug. 2006    rev 1.0
       original version

   hm  25. oct. 2008   rev 1.1
       optimized code

   hm  14. mar. 2009   rev 1.2
       removed double assignments

   *)
END_FUNCTION_BLOCK

FUNCTION_BLOCK "SHR_8PLE"   // FB89, SCL
TITLE = SHR_8PLE
{ S7_Optimized_Access := 'FALSE' }
AUTHOR : hugo
FAMILY : FFETRIG
NAME : SHR8PLE
VERSION : 1.0
// 8 bit shift register with reset and parallel load
// the register can shift up or down
// it also has a serial input.
// the Din input is on Bit0 for up shift and on bit 7 for down shift
// the Dout output is on Bit7 for up shift and on bit 0 for down shift
// paralle clock is performed clock synchron while a shift is performed first and then the register is reloaded
   VAR_INPUT
      Din : Bool;
      Dload : Byte;
      CLK : Bool;
      UP : Bool := TRUE;
      load : Bool;
      RST : Bool;
   END_VAR
   VAR_OUTPUT
      DOut : Bool;
   END_VAR
   VAR
      edge : Bool := TRUE;
      register : Byte;
      tregister AT register : Array[0..7] of Bool;
   END_VAR
BEGIN


     (* flankenerkennung clk wird high und edge war high reset ist nicht aktiv und set ist nicht aktiv *)
     IF #CLK AND #edge AND NOT #RST THEN
         #edge := FALSE;  (* flanke wurde erkannt und weitere flankenerkennung wird verhindert bis edge wieder true ist *)
         (* hier ist der code für das flankenevent *)
         IF #UP THEN                      (*shift up *)
             #register := SHL(IN:=#register,N:=1);
             #tregister[0] := #Din;
             #DOut := #tregister[7];
         ELSE                                (* shift down *);
             #register := SHR(IN:=#register,N:=1);
             #tregister[7] := #Din;
             #DOut := #tregister[0];
         END_IF;
         IF #load THEN                            (* the byte on Din will be loaded if load = true *)
             #register := #Dload;
             IF #UP THEN #DOut := #tregister[7]; ELSE #DOut := #tregister[0]; END_IF;
         END_IF;
     END_IF;
     IF NOT #CLK THEN #edge := TRUE; END_IF;  (* sobald clk wieder low wird warten auf nächste flanke *)
     IF #RST THEN                                 (* wenn reset aktiv dann ausgang rücksetzen *)
         #register := 0;
         #DOut := FALSE;
     END_IF;
END_FUNCTION_BLOCK

FUNCTION_BLOCK "SHR_8UDE"   // FB90, SCL
TITLE = SHR_8UDE
{ S7_Optimized_Access := 'FALSE' }
AUTHOR : hugo
FAMILY : FFETRIG
NAME : SHR8UDE
VERSION : 1.2
// 8 bit shift register with reset
   VAR_INPUT
      SET : Bool;
      D0 : Bool;
      D7 : Bool;
      CLK : Bool;
      DN : Bool;
      RST : Bool;
   END_VAR
   VAR_OUTPUT
      Q0 : Bool;
      Q1 : Bool;
      Q2 : Bool;
      Q3 : Bool;
      Q4 : Bool;
      Q5 : Bool;
      Q6 : Bool;
      Q7 : Bool;
   END_VAR
   VAR
      "m" : Bool;
   END_VAR
BEGIN


   (* trig.Q signals a rising edge on clk *)
   (* trig(clk := clk); *)

   IF #SET OR #RST THEN
       #Q0 := NOT #RST;
       #Q1 := #Q0;
       #Q2 := #Q0;
       #Q3 := #Q0;
       #Q4 := #Q0;
       #Q5 := #Q0;
       #Q6 := #Q0;
       #Q7 := #Q0;
   ELSIF #CLK AND NOT #"m" THEN
       IF #DN THEN
           #Q0 := #Q1;
           #Q1 := #Q2;
           #Q2 := #Q3;
           #Q3 := #Q4;
           #Q4 := #Q5;
           #Q5 := #Q6;
           #Q6 := #Q7;
           #Q7 := #D7;
       ELSE
           #Q7 := #Q6;
           #Q6 := #Q5;
           #Q5 := #Q4;
           #Q4 := #Q3;
           #Q3 := #Q2;
           #Q2 := #Q1;
           #Q1 := #Q0;
           #Q0 := #D0;
       END_IF;
   END_IF;

   #"m" := #CLK;


   (* revision history
   hm  4. aug. 2006    rev 1.0
       original version

   hm  25. oct. 2008   rev 1.1
       optimized code

   hm  14. mar. 2009   rev 1.2
       removed double assignments

   *)
END_FUNCTION_BLOCK

FUNCTION_BLOCK "TOGGLE"   // FB92, SCL
TITLE = TOGGLE
{ S7_Optimized_Access := 'FALSE' }
AUTHOR : hugo
FAMILY : FFETRIG
NAME : TOGGLE
VERSION : 1.1
// toggle flip flop the output changes state with every rising edge of clk.
   VAR_INPUT
      CLK : Bool;
      rst : Bool;
   END_VAR
   VAR_OUTPUT
      Q : Bool;
   END_VAR
   VAR
      edge : Bool;
   END_VAR
BEGIN


   IF #rst THEN
       #Q := 0;
   ELSIF #CLK AND NOT #edge THEN
       #Q := NOT #Q;
   END_IF;
   #edge := #CLK;


   (* revision history

   hm  13.9.2007       rev 1.0
       original version

   hm  30. oct. 2008   rev 1.1
       deleted unnecessary init

   *)
END_FUNCTION_BLOCK

FUNCTION "INC" : Int   // FC90, SCL
TITLE = INC
{ S7_Optimized_Access := 'FALSE' }
AUTHOR : hugo
FAMILY : MATH
NAME : INC
VERSION : 1.1
// This is a increment function which increments the input X by the value D and compares the result with M.
// if the output exceeds M it will continue to count from 0 again.
   VAR_INPUT
      X : Int;
      D : Int;
      "M" : Int;
   END_VAR
BEGIN


     #INC := (#X + #D + #"M" + 1) MOD (#"M" + 1);

   (* revision history
   hm  7. feb 2007   REV 1.0
     original version

   hm  15. jan 2008  rev 1.1
     allow for neagtive increment

   *)
END_FUNCTION

// ===== PLC "Logic FF pulse triggered"  Unspecific CPU S7 300 =====

FUNCTION_BLOCK "LTCH"   // FB85, SCL
TITLE = LTCH
{ S7_Optimized_Access := 'FALSE' }
AUTHOR : hugo
FAMILY : FFPTRIG
NAME : LTCH
VERSION : 1.2
// Transparent Latch with asynchronous reset
   VAR_INPUT
      D : Bool;
      L : Bool;
      RST : Bool;
   END_VAR
   VAR_OUTPUT
      Q : Bool;
   END_VAR
BEGIN


   (* as long as L is true, the latch is transparent and and change of D is transferred to Q *)
   (* of course only when there is no asynchronous reset *)
   IF #RST THEN       (* if asynchronous reset then Q=0 *)
       #Q := FALSE;
   ELSIF #L THEN      (* latch is transparent *)
       #Q := #D;
   END_IF;


   (* revision history
   hm  4. aug 2006     rev 1.0
       original version

   hm  27. dec 2007    rev 1.1
       changed code for better performance

   hm  30. oct. 2008   rev 1.2
       deleted unnecessary init with 0

   *)
END_FUNCTION_BLOCK

FUNCTION_BLOCK "LTCH_4"   // FB86, SCL
TITLE = LTCH_4
{ S7_Optimized_Access := 'FALSE' }
AUTHOR : hugo
FAMILY : FFPTRIG
NAME : LTCH_4
VERSION : 1.3
// Quad Transparent Latch with asynchronous reset
   VAR_INPUT
      D0 : Bool;
      D1 : Bool;
      D2 : Bool;
      D3 : Bool;
      L : Bool;
      RST : Bool;
   END_VAR
   VAR_OUTPUT
      Q0 : Bool;
      Q1 : Bool;
      Q2 : Bool;
      Q3 : Bool;
   END_VAR
BEGIN


   (* as long as L is true, the latch is transparent and and change of D is transferred to Q *)
   (* of course only when there is no asynchronous reset *)
   IF #RST THEN       (* if asynchronous reset then Q=0 *)
       #Q0 := FALSE;
       #Q1 := FALSE;
       #Q2 := FALSE;
       #Q3 := FALSE;
   ELSIF #L THEN      (* latch is transparent *)
       #Q0 := #D0;
       #Q1 := #D1;
       #Q2 := #D2;
       #Q3 := #D3;
   END_IF;


   (* revision history
   hm  4. aug 2006 rev 1.0
       original version

   hm  27. dec 2007    rev 1.1
       changed code for better performance

   hm  30. oct. 2008   rev 1.2
       deleted unnecessary init with 0

   hm  14. mar. 2009   rev 1.3
       removed double assignments

   *)
END_FUNCTION_BLOCK

FUNCTION_BLOCK "STORE_8"   // FB91, SCL
TITLE = STORE_8
{ S7_Optimized_Access := 'FALSE' }
AUTHOR : hugo
FAMILY : FFETRIG
NAME : STORE_8
VERSION : 1.2
// Store_4 stores up to 4 boolean inputs until a reset is clearing the outputs.
// the respective output is set with a true at the respective input and stays true until a reset is generated.
// a set input is used to set all outputs true at the same time, independent of their inputs.
// a clear input is used to reset only the lowest priority of the outputs one at a time.
// the lowest priority is q3.
   VAR_INPUT
      Set : Bool;
      D0 : Bool;
      D1 : Bool;
      D2 : Bool;
      D3 : Bool;
      D4 : Bool;
      D5 : Bool;
      D6 : Bool;
      D7 : Bool;
      Clr : Bool;
      Rst : Bool;
   END_VAR
   VAR_OUTPUT
      Q0 : Bool;
      Q1 : Bool;
      Q2 : Bool;
      Q3 : Bool;
      Q4 : Bool;
      Q5 : Bool;
      Q6 : Bool;
      Q7 : Bool;
   END_VAR
   VAR
      edge : Bool;
   END_VAR
BEGIN


   IF #Rst OR #Set THEN
       #Q0 := NOT #Rst;
       #Q1 := #Q0;
       #Q2 := #Q0;
       #Q3 := #Q0;
       #Q4 := #Q0;
       #Q5 := #Q0;
       #Q6 := #Q0;
       #Q7 := #Q0;
   ELSE
       IF #D0 THEN #Q0 := TRUE; END_IF;
       IF #D1 THEN #Q1 := TRUE; END_IF;
       IF #D2 THEN #Q2 := TRUE; END_IF;
       IF #D3 THEN #Q3 := TRUE; END_IF;
       IF #D4 THEN #Q4 := TRUE; END_IF;
       IF #D5 THEN #Q5 := TRUE; END_IF;
       IF #D6 THEN #Q6 := TRUE; END_IF;
       IF #D7 THEN #Q7 := TRUE; END_IF;

